   IOField "I/O field_31" at 476,376 size 58x21; FormatPattern s99999
      ProcessValue <- "AIx_DB_Flow_4_SP_SC"
   IOField "I/O field_32" at 250,358 size 58x21; FormatPattern 99999
      ProcessValue <- "AIx_DB_Flow_4_SP_HH"
   IOField "I/O field_33" at 250,378 size 58x21; FormatPattern 99999
      ProcessValue <- "AIx_DB_Flow_4_SP_H"
   IOField "I/O field_34" at 250,398 size 58x21; FormatPattern s99999
      ProcessValue <- "AIx_DB_Flow_4_SP_L"
   IOField "I/O field_35" at 250,418 size 58x21; FormatPattern s99999
      ProcessValue <- "AIx_DB_Flow_4_SP_LL"
   IOField "I/O field_36" at 550,356 size 58x21; FormatPattern 999
      ProcessValue <- "AIx_DB_Flow_4_Timers_NC_SP"
   IOField "I/O field_37" at 550,376 size 58x21; FormatPattern 999
      ProcessValue <- "AIx_DB_Flow_4_Timers_SC_SP"
   IOField "I/O field_38" at 324,358 size 58x21; FormatPattern 999
      ProcessValue <- "AIx_DB_Flow_4_Timers_HH_SP"
   IOField "I/O field_39" at 324,378 size 58x21; FormatPattern 999
      ProcessValue <- "AIx_DB_Flow_4_Timers_H_SP"
   IOField "I/O field_40" at 324,398 size 58x21; FormatPattern 999
      ProcessValue <- "AIx_DB_Flow_4_Timers_L_SP"
   IOField "I/O field_41" at 324,418 size 58x21; FormatPattern 999
      ProcessValue <- "AIx_DB_Flow_4_Timers_LL_SP"
   IOField "I/O field_42" at 586,326 size 65x25; FormatPattern s99999
      ProcessValue <- "AIx_DB_Flow_4_Signal"
   TextField "Text field_29" at 214,330 size 68x22; Text 'Уставка'
   TextField "Text field_30" at 303,330 size 79x22; Text 'Время (с)'
   Button "Button_1" at 7,5 size 96x32; TextOff 'Насосы'; Authorization "Admin"
      on Release: ActivateScreen("Dos", 0); SetTag("settings", 1)
      Appearance <- "settings"
   Button "Button_2" at 7,51 size 96x32; TextOff 'Расход-1'; Authorization "Admin"
      on Release: ActivateScreen("Flow", 0); SetTag("settings", 2)
      Appearance <- "settings"
   Button "Button_3" at 7,140 size 96x32; TextOff 'Мутность'; Authorization "Admin"
      on Release: ActivateScreen("Trans", 0); SetTag("settings", 4)
      Appearance <- "settings"
   Button "Button_5" at 7,184 size 96x32; TextOff 'DI'; Authorization "Admin"
      on Release: ActivateScreen("DI", 0); SetTag("settings", 5)
      Appearance <- "settings"
   Button "Button_6" at 7,229 size 96x32; TextOff 'DO'; Authorization "Admin"
      on Release: ActivateScreen("DO", 0); SetTag("settings", 6)
      Appearance <- "settings"
   Button "Button_4" at 7,274 size 96x32; TextOff 'PID'; Authorization "Admin"
      on Release: ActivateScreen("PID_settings", 0); SetTag("settings", 7)
      Appearance <- "settings"
   Button "Button_15" at 7,95 size 96x32; TextOff 'Расход-2'; Authorization "Admin"
      on Release: ActivateScreen("Flow_1", 0); SetTag("settings", 3)
      Appearance <- "settings"
*)

(* ===== HMI "HMI_RT_4" =====
system functions are stored by id; their names below are inferred from use
connection "HMI_Connection_2": ETHERNET, SMART_S7_1200_OMS

HMI tags "Default tag table"
   "Comm_1_DB_Mix_3_Status" : Int = PLC Comm_1_DB.Mix_3_Status AT %DB11.DBW24, 1 s
   "Comm_1_DB_Mix_2_Status" : Int = PLC Comm_1_DB.Mix_2_Status AT %DB11.DBW18, 1 s
   "Comm_1_DB_Mix_1_Status" : Int = PLC Comm_1_DB.Mix_1_Status AT %DB11.DBW12, 1 s
   "Comm_1_DB_Level" : Real = PLC Comm_1_DB.Level AT %DB11.DBD38, 1 s
   "Comm_2_DB_Level" : Real = PLC Comm_2_DB.Level AT %DB12.DBD38, 1 s
   "Comm_2_DB_Mix_1_Status" : Int = PLC Comm_2_DB.Mix_1_Status AT %DB12.DBW12, 1 s
   "Comm_2_DB_Mix_2_Status" : Int = PLC Comm_2_DB.Mix_2_Status AT %DB12.DBW18, 1 s
   "Comm_2_DB_Mix_3_Status" : Int = PLC Comm_2_DB.Mix_3_Status AT %DB12.DBW24, 1 s
   "Any_Hand" : Bool = PLC Any_Hand AT %M5.0, 1 s
   "Logick_DB_Start" : Bool = PLC Logick_DB.Start AT %DB1.DBX0.0, 1 s
   "Logick_DB_Hand" : Bool = PLC Logick_DB.Hand AT %DB1.DBX0.1, 1 s
   "Logick_DB_Use_M1" : Bool = PLC Logick_DB.Use_M1 AT %DB1.DBX0.6, 1 s
   "Logick_DB_Use_M3" : Bool = PLC Logick_DB.Use_M3 AT %DB1.DBX1.0, 1 s
   "Logick_DB_REQ_M2_1" : Bool = PLC Logick_DB.REQ_M2_1 AT %DB1.DBX1.3, 1 s
   "Logick_DB_Res_M1" : Bool = PLC Logick_DB.Res_M1 AT %DB1.DBX1.1, 1 s
   "Logick_DB_Res_M3" : Bool = PLC Logick_DB.Res_M3 AT %DB1.DBX1.2, 1 s
   "RS232_DB_Mass_1" : Real = PLC RS232_DB.Mass_1 AT %DB2.DBD0, 1 s
   "Statistics_DB_Today_1" : Real = PLC Statistics_DB.Today_1 AT %DB4.DBD40, 1 s
   "Statistics_DB_Mass_2" : Real = PLC Statistics_DB.Mass_2 AT %DB4.DBD4, 1 s
   "Statistics_DB_Mass_1" : Real = PLC Statistics_DB.Mass_1 AT %DB4.DBD0, 1 s
   "Statistics_DB_Today_2" : Real = PLC Statistics_DB.Today_2 AT %DB4.DBD44, 1 s
   "Logick_DB_Fix_1" : Bool = PLC Logick_DB.Fix_1 AT %DB1.DBX0.2, 1 s
   "Logick_DB_Fix_D_1" : Real = PLC Logick_DB.Fix_D_1 AT %DB1.DBD48, 1 s
   "Logick_DB_D_1" : Real = PLC Logick_DB.D_1 AT %DB1.DBD56, 1 s
   "Logick_DB_Fix_2" : Bool = PLC Logick_DB.Fix_2 AT %DB1.DBX0.3, 1 s
   "Logick_DB_Fix_D_2" : Real = PLC Logick_DB.Fix_D_2 AT %DB1.DBD52, 1 s
   "Logick_DB_D_2" : Real = PLC Logick_DB.D_2 AT %DB1.DBD60, 1 s
   "Comm_1_DB_Warning" : Bool = PLC Comm_1_DB.Warning AT %DB11.DBX48.2, 1 s
   "Comm_2_DB_Warning" : Bool = PLC Comm_2_DB.Warning AT %DB12.DBX48.2, 1 s
   "Logick_DB_C_1" : Real = PLC Logick_DB.C_1 AT %DB1.DBD64, 1 s
   "Logick_DB_C_2" : Real = PLC Logick_DB.C_2 AT %DB1.DBD68, 1 s
   "Statistics_DB_Zero_1" : Real = PLC Statistics_DB.Zero_1 AT %DB4.DBD64, 1 s
   "RS232_DB_Mass_2" : Real = PLC RS232_DB.Mass_2 AT %DB2.DBD4, 1 s
   "Statistics_DB_Zero_2" : Real = PLC Statistics_DB.Zero_2 AT %DB4.DBD68, 1 s
   "Statistics_DB_Last_1" : Real = PLC Statistics_DB.Last_1 AT %DB4.DBD24, 1 s
   "Statistics_DB_Delta_1" : Real = PLC Statistics_DB.Delta_1 AT %DB4.DBD32, 1 s
   "Statistics_DB_Max_D_1" : Real = PLC Statistics_DB.Max_D_1 AT %DB4.DBD16, 1 s
   "Statistics_DB_Min_D_1" : Real = PLC Statistics_DB.Min_D_1 AT %DB4.DBD8, 1 s
   "Statistics_DB_T_SP_M" : Int = PLC Statistics_DB.T.SP_M AT %DB4.DBW580, 1 s
   "Statistics_DB_T_SP_S" : Int = PLC Statistics_DB.T.SP_S AT %DB4.DBW582, 1 s
   "Sync" : Bool = PLC Sync_1 AT %M10.0, 1 s
   "Sync_2" : Bool = PLC Sync_2 AT %M10.1, 1 s
   "Statistics_DB_Delta_2" : Real = PLC Statistics_DB.Delta_2 AT %DB4.DBD36, 1 s
   "Statistics_DB_Last_2" : Real = PLC Statistics_DB.Last_2 AT %DB4.DBD28, 1 s
   "Statistics_DB_Max_D_2" : Real = PLC Statistics_DB.Max_D_2 AT %DB4.DBD20, 1 s
   "Statistics_DB_Min_D_2" : Real = PLC Statistics_DB.Min_D_2 AT %DB4.DBD12, 1 s
   "DIx_DB_Heat_4_Signal" : Bool = PLC DIx_DB.Heat_4.Signal AT %DB200.DBX122.0, 1 s
   "DIx_DB_Heat_4_Input" : Bool = PLC DIx_DB.Heat_4.Input AT %DB200.DBX120.0, 1 s
   "DIx_DB_Heat_1_Inverse" : Bool = PLC DIx_DB.Heat_1.Inverse AT %DB200.DBX64.3, 1 s
   "Any_Alm" : Bool = PLC Any_Alm AT %M6.0, 1 s
   "Statistics_DB_Today_Int" : Int = PLC Statistics_DB.Today_Int AT %DB4.DBW74, 1 s
   "Time_Save" : Bool = PLC "Time".Save AT %DB13.DBX38.0, 1 s
   "Time_Year" : UInt = PLC "Time".Year AT %DB13.DBW28, 1 s
   "Time_Month" : UInt = PLC "Time".Month AT %DB13.DBW30, 1 s
   "Time_Day" : UInt = PLC "Time".Day AT %DB13.DBW32, 1 s
   "Time_Hour" : UInt = PLC "Time".Hour AT %DB13.DBW34, 1 s
   "Time_Minutes" : UInt = PLC "Time".Minutes AT %DB13.DBW36, 1 s
   "Time_Today_YEAR" : UInt = PLC "Time".Today.YEAR AT %DB13.DBW0, 1 s
   "Time_Today_MONTH" : USInt = PLC "Time".Today.MONTH AT %DB13.DBB2, 1 s
   "Time_Today_DAY" : USInt = PLC "Time".Today.DAY AT %DB13.DBB3, 1 s
   "Time_Today_WEEKDAY" : USInt = PLC "Time".Today.WEEKDAY AT %DB13.DBB4, 1 s
   "Time_Today_HOUR" : USInt = PLC "Time".Today.HOUR AT %DB13.DBB5, 1 s
   "Time_Today_MINUTE" : USInt = PLC "Time".Today.MINUTE AT %DB13.DBB6, 1 s
   "Reset_All" : Bool = PLC Reset_All AT %M3.1, 1 s
   "Logick_DB_Low_REQ" : Bool = PLC Logick_DB.Low_REQ AT %DB1.DBX2.0, 1 s
   "Logick_DB_Low_view" : Bool = PLC Logick_DB.Low_view AT %DB1.DBX2.2, 1 s
   "Logick_DB_Low_SP_M" : Int = PLC Logick_DB.Low.SP_M AT %DB1.DBW72, 1 s
   "Logick_DB_Low_CMD" : Bool = PLC Logick_DB.Low_CMD AT %DB1.DBX2.1, 1 s
   "Logick_DB_Max_SP" : Real = PLC Logick_DB.Max_SP AT %DB1.DBD36, 1 s
   "Logick_DB_Min_SP" : Real = PLC Logick_DB.Min_SP AT %DB1.DBD32, 1 s
   "Logick_DB_Low_use" : Bool = PLC Logick_DB.Low_use AT %DB1.DBX1.7, 1 s

HMI tags "HMI"
   "settings" : Int, internal

HMI tags "xDI"
   "DIx_DB_M1_QF_Input" : Bool = PLC DIx_DB.M1_QF.Input AT %DB200.DBX0.0, 1 s
   "DIx_DB_M1_QF_Signal" : Bool = PLC DIx_DB.M1_QF.Signal AT %DB200.DBX2.0, 1 s
   "DIx_DB_M1_QF_Hand" : Bool = PLC DIx_DB.M1_QF.Hand AT %DB200.DBX4.0, 1 s
   "DIx_DB_M1_QF_Start_M" : Bool = PLC DIx_DB.M1_QF.Start_M AT %DB200.DBX4.1, 1 s
   "DIx_DB_M1_QF_Inverse" : Bool = PLC DIx_DB.M1_QF.Inverse AT %DB200.DBX4.3, 1 s
   "DIx_DB_M1_QF_Filter_On_SP" : Int = PLC DIx_DB.M1_QF.Filter_On.SP AT %DB200.DBW6, 1 s
   "DIx_DB_M1_QF_Filter_Off_SP" : Int = PLC DIx_DB.M1_QF.Filter_Off.SP AT %DB200.DBW12, 1 s
   "DIx_DB_M2_QF_Input" : Bool = PLC DIx_DB.M2_QF.Input AT %DB200.DBX20.0, 1 s
   "DIx_DB_M2_QF_Signal" : Bool = PLC DIx_DB.M2_QF.Signal AT %DB200.DBX22.0, 1 s
   "DIx_DB_M2_QF_Hand" : Bool = PLC DIx_DB.M2_QF.Hand AT %DB200.DBX24.0, 1 s
   "DIx_DB_M2_QF_Start_M" : Bool = PLC DIx_DB.M2_QF.Start_M AT %DB200.DBX24.1, 1 s
   "DIx_DB_M2_QF_Inverse" : Bool = PLC DIx_DB.M2_QF.Inverse AT %DB200.DBX24.3, 1 s
   "DIx_DB_M2_QF_Filter_On_SP" : Int = PLC DIx_DB.M2_QF.Filter_On.SP AT %DB200.DBW26, 1 s
   "DIx_DB_M2_QF_Filter_Off_SP" : Int = PLC DIx_DB.M2_QF.Filter_Off.SP AT %DB200.DBW32, 1 s
   "DIx_DB_M3_QF_Input" : Bool = PLC DIx_DB.M3_QF.Input AT %DB200.DBX40.0, 1 s
   "DIx_DB_M3_QF_Signal" : Bool = PLC DIx_DB.M3_QF.Signal AT %DB200.DBX42.0, 1 s
   "DIx_DB_M3_QF_Hand" : Bool = PLC DIx_DB.M3_QF.Hand AT %DB200.DBX44.0, 1 s
   "DIx_DB_M3_QF_Start_M" : Bool = PLC DIx_DB.M3_QF.Start_M AT %DB200.DBX44.1, 1 s
   "DIx_DB_M3_QF_Inverse" : Bool = PLC DIx_DB.M3_QF.Inverse AT %DB200.DBX44.3, 1 s
   "DIx_DB_M3_QF_Filter_On_SP" : Int = PLC DIx_DB.M3_QF.Filter_On.SP AT %DB200.DBW46, 1 s
   "DIx_DB_M3_QF_Filter_Off_SP" : Int = PLC DIx_DB.M3_QF.Filter_Off.SP AT %DB200.DBW52, 1 s
   "DIx_DB_Heat_1_Input" : Bool = PLC DIx_DB.Heat_1.Input AT %DB200.DBX60.0, 1 s
   "DIx_DB_Heat_1_Signal" : Bool = PLC DIx_DB.Heat_1.Signal AT %DB200.DBX62.0, 1 s
   "DIx_DB_Heat_1_Hand" : Bool = PLC DIx_DB.Heat_1.Hand AT %DB200.DBX64.0, 1 s
   "DIx_DB_Heat_1_Start_M" : Bool = PLC DIx_DB.Heat_1.Start_M AT %DB200.DBX64.1, 1 s
   "DIx_DB_Heat_1_Filter_On_SP" : Int = PLC DIx_DB.Heat_1.Filter_On.SP AT %DB200.DBW66, 1 s
   "DIx_DB_Heat_1_Filter_Off_SP" : Int = PLC DIx_DB.Heat_1.Filter_Off.SP AT %DB200.DBW72, 1 s
   "DIx_DB_Heat_2_Filter_Off_SP" : Int = PLC DIx_DB.Heat_2.Filter_Off.SP AT %DB200.DBW92, 1 s
   "DIx_DB_Heat_2_Filter_On_SP" : Int = PLC DIx_DB.Heat_2.Filter_On.SP AT %DB200.DBW86, 1 s
   "DIx_DB_Heat_2_Inverse" : Bool = PLC DIx_DB.Heat_2.Inverse AT %DB200.DBX84.3, 1 s
   "DIx_DB_Heat_2_Start_M" : Bool = PLC DIx_DB.Heat_2.Start_M AT %DB200.DBX84.1, 1 s
   "DIx_DB_Heat_2_Hand" : Bool = PLC DIx_DB.Heat_2.Hand AT %DB200.DBX84.0, 1 s
   "DIx_DB_Heat_2_Signal" : Bool = PLC DIx_DB.Heat_2.Signal AT %DB200.DBX82.0, 1 s
   "DIx_DB_Heat_2_Input" : Bool = PLC DIx_DB.Heat_2.Input AT %DB200.DBX80.0, 1 s
   "DIx_DB_Heat_3_Input" : Bool = PLC DIx_DB.Heat_3.Input AT %DB200.DBX100.0, 1 s
   "DIx_DB_Heat_3_Signal" : Bool = PLC DIx_DB.Heat_3.Signal AT %DB200.DBX102.0, 1 s
   "DIx_DB_Heat_3_Hand" : Bool = PLC DIx_DB.Heat_3.Hand AT %DB200.DBX104.0, 1 s
   "DIx_DB_Heat_3_Start_M" : Bool = PLC DIx_DB.Heat_3.Start_M AT %DB200.DBX104.1, 1 s
   "DIx_DB_Heat_3_Inverse" : Bool = PLC DIx_DB.Heat_3.Inverse AT %DB200.DBX104.3, 1 s
   "DIx_DB_Heat_3_Filter_Off_SP" : Int = PLC DIx_DB.Heat_3.Filter_Off.SP AT %DB200.DBW112, 1 s
   "DIx_DB_Heat_3_Filter_On_SP" : Int = PLC DIx_DB.Heat_3.Filter_On.SP AT %DB200.DBW106, 1 s
   "DIx_DB_AllBlock_Input" : Bool = PLC DIx_DB.AllBlock.Input AT %DB200.DBX140.0, 1 s
   "DIx_DB_AllBlock_Signal" : Bool = PLC DIx_DB.AllBlock.Signal AT %DB200.DBX142.0, 1 s
   "DIx_DB_AllBlock_Hand" : Bool = PLC DIx_DB.AllBlock.Hand AT %DB200.DBX144.0, 1 s
   "DIx_DB_AllBlock_Start_M" : Bool = PLC DIx_DB.AllBlock.Start_M AT %DB200.DBX144.1, 1 s
   "DIx_DB_AllBlock_Inverse" : Bool = PLC DIx_DB.AllBlock.Inverse AT %DB200.DBX144.3, 1 s
   "DIx_DB_AllBlock_Filter_On_SP" : Int = PLC DIx_DB.AllBlock.Filter_On.SP AT %DB200.DBW146, 1 s
   "DIx_DB_AllBlock_Filter_Off_SP" : Int = PLC DIx_DB.AllBlock.Filter_Off.SP AT %DB200.DBW152, 1 s
   "DIx_DB_Mass_1_Input" : Bool = PLC DIx_DB.Mass_1.Input AT %DB200.DBX160.0, 1 s
   "DIx_DB_Mass_1_Signal" : Bool = PLC DIx_DB.Mass_1.Signal AT %DB200.DBX162.0, 1 s
   "DIx_DB_Mass_1_Hand" : Bool = PLC DIx_DB.Mass_1.Hand AT %DB200.DBX164.0, 1 s
   "DIx_DB_Mass_1_Start_M" : Bool = PLC DIx_DB.Mass_1.Start_M AT %DB200.DBX164.1, 1 s
   "DIx_DB_Mass_1_Inverse" : Bool = PLC DIx_DB.Mass_1.Inverse AT %DB200.DBX164.3, 1 s
   "DIx_DB_Mass_1_Filter_On_SP" : Int = PLC DIx_DB.Mass_1.Filter_On.SP AT %DB200.DBW166, 1 s
   "DIx_DB_Mass_1_Filter_Off_SP" : Int = PLC DIx_DB.Mass_1.Filter_Off.SP AT %DB200.DBW172, 1 s
   "DIx_DB_Mass_2_Input" : Bool = PLC DIx_DB.Mass_2.Input AT %DB200.DBX180.0, 1 s
   "DIx_DB_Mass_2_Signal" : Bool = PLC DIx_DB.Mass_2.Signal AT %DB200.DBX182.0, 1 s
   "DIx_DB_Mass_2_Hand" : Bool = PLC DIx_DB.Mass_2.Hand AT %DB200.DBX184.0, 1 s
   "DIx_DB_Mass_2_Start_M" : Bool = PLC DIx_DB.Mass_2.Start_M AT %DB200.DBX184.1, 1 s
   "DIx_DB_Mass_2_Inverse" : Bool = PLC DIx_DB.Mass_2.Inverse AT %DB200.DBX184.3, 1 s
   "DIx_DB_Mass_2_Filter_On_SP" : Int = PLC DIx_DB.Mass_2.Filter_On.SP AT %DB200.DBW186, 1 s
   "DIx_DB_Mass_2_Filter_Off_SP" : Int = PLC DIx_DB.Mass_2.Filter_Off.SP AT %DB200.DBW192, 1 s
   "DIx_DB_Heat_4_Hand" : Bool = PLC DIx_DB.Heat_4.Hand AT %DB200.DBX124.0, 1 s
   "DIx_DB_Heat_4_Start_M" : Bool = PLC DIx_DB.Heat_4.Start_M AT %DB200.DBX124.1, 1 s
   "DIx_DB_Heat_4_Inverse" : Bool = PLC DIx_DB.Heat_4.Inverse AT %DB200.DBX124.3, 1 s
   "DIx_DB_Heat_4_Filter_On_SP" : Int = PLC DIx_DB.Heat_4.Filter_On.SP AT %DB200.DBW126, 1 s
   "DIx_DB_Heat_4_Filter_Off_SP" : Int = PLC DIx_DB.Heat_4.Filter_Off.SP AT %DB200.DBW132, 1 s

HMI tags "xDO"
   "DOx_DB_M1_CMD_Start_A" : Bool = PLC DOx_DB.M1_CMD.Start_A AT %DB201.DBX0.0, 1 s
   "DOx_DB_M1_CMD_Q" : Bool = PLC DOx_DB.M1_CMD.Q AT %DB201.DBX0.2, 1 s
   "DOx_DB_M1_CMD_Hand" : Bool = PLC DOx_DB.M1_CMD.Hand AT %DB201.DBX2.0, 1 s
   "DOx_DB_M1_CMD_Start_M" : Bool = PLC DOx_DB.M1_CMD.Start_M AT %DB201.DBX2.1, 1 s
   "DOx_DB_M1_CMD_Simulation" : Bool = PLC DOx_DB.M1_CMD.Simulation AT %DB201.DBX2.2, 1 s
   "DOx_DB_M1_CMD_Inverse" : Bool = PLC DOx_DB.M1_CMD.Inverse AT %DB201.DBX2.3, 1 s
   "DOx_DB_M2_CMD_Start_A" : Bool = PLC DOx_DB.M2_CMD.Start_A AT %DB201.DBX10.0, 1 s
   "DOx_DB_M2_CMD_Q" : Bool = PLC DOx_DB.M2_CMD.Q AT %DB201.DBX10.2, 1 s
   "DOx_DB_M2_CMD_Hand" : Bool = PLC DOx_DB.M2_CMD.Hand AT %DB201.DBX12.0, 1 s
   "DOx_DB_M2_CMD_Start_M" : Bool = PLC DOx_DB.M2_CMD.Start_M AT %DB201.DBX12.1, 1 s
   "DOx_DB_M2_CMD_Simulation" : Bool = PLC DOx_DB.M2_CMD.Simulation AT %DB201.DBX12.2, 1 s
   "DOx_DB_M2_CMD_Inverse" : Bool = PLC DOx_DB.M2_CMD.Inverse AT %DB201.DBX12.3, 1 s
   "DOx_DB_M3_CMD_Start_A" : Bool = PLC DOx_DB.M3_CMD.Start_A AT %DB201.DBX20.0, 1 s
   "DOx_DB_M3_CMD_Q" : Bool = PLC DOx_DB.M3_CMD.Q AT %DB201.DBX20.2, 1 s
   "DOx_DB_M3_CMD_Hand" : Bool = PLC DOx_DB.M3_CMD.Hand AT %DB201.DBX22.0, 1 s
   "DOx_DB_M3_CMD_Start_M" : Bool = PLC DOx_DB.M3_CMD.Start_M AT %DB201.DBX22.1, 1 s
   "DOx_DB_M3_CMD_Simulation" : Bool = PLC DOx_DB.M3_CMD.Simulation AT %DB201.DBX22.2, 1 s
   "DOx_DB_M3_CMD_Inverse" : Bool = PLC DOx_DB.M3_CMD.Inverse AT %DB201.DBX22.3, 1 s
   "DOx_DB_LED_Error_1_Start_A" : Bool = PLC DOx_DB.LED_Error_1.Start_A AT %DB201.DBX30.0, 1 s
   "DOx_DB_LED_Error_1_Q" : Bool = PLC DOx_DB.LED_Error_1.Q AT %DB201.DBX30.2, 1 s
   "DOx_DB_LED_Error_1_Hand" : Bool = PLC DOx_DB.LED_Error_1.Hand AT %DB201.DBX32.0, 1 s
   "DOx_DB_LED_Error_1_Simulation" : Bool = PLC DOx_DB.LED_Error_1.Simulation AT %DB201.DBX32.2, 1 s
   "DOx_DB_LED_Error_1_Start_M" : Bool = PLC DOx_DB.LED_Error_1.Start_M AT %DB201.DBX32.1, 1 s
   "DOx_DB_LED_Error_1_Inverse" : Bool = PLC DOx_DB.LED_Error_1.Inverse AT %DB201.DBX32.3, 1 s
   "DOx_DB_LED_Error_2_Start_A" : Bool = PLC DOx_DB.LED_Error_2.Start_A AT %DB201.DBX40.0, 1 s
   "DOx_DB_LED_Error_2_Q" : Bool = PLC DOx_DB.LED_Error_2.Q AT %DB201.DBX40.2, 1 s
   "DOx_DB_LED_Error_2_Hand" : Bool = PLC DOx_DB.LED_Error_2.Hand AT %DB201.DBX42.0, 1 s
   "DOx_DB_LED_Error_2_Start_M" : Bool = PLC DOx_DB.LED_Error_2.Start_M AT %DB201.DBX42.1, 1 s
   "DOx_DB_LED_Error_2_Simulation" : Bool = PLC DOx_DB.LED_Error_2.Simulation AT %DB201.DBX42.2, 1 s
   "DOx_DB_LED_Error_2_Inverse" : Bool = PLC DOx_DB.LED_Error_2.Inverse AT %DB201.DBX42.3, 1 s
   "DOx_DB_LED_Alarm_Start_A" : Bool = PLC DOx_DB.LED_Alarm.Start_A AT %DB201.DBX50.0, 1 s
   "DOx_DB_LED_Alarm_Q" : Bool = PLC DOx_DB.LED_Alarm.Q AT %DB201.DBX50.2, 1 s
   "DOx_DB_LED_Alarm_Hand" : Bool = PLC DOx_DB.LED_Alarm.Hand AT %DB201.DBX52.0, 1 s
   "DOx_DB_LED_Alarm_Start_M" : Bool = PLC DOx_DB.LED_Alarm.Start_M AT %DB201.DBX52.1, 1 s
   "DOx_DB_LED_Alarm_Simulation" : Bool = PLC DOx_DB.LED_Alarm.Simulation AT %DB201.DBX52.2, 1 s
   "DOx_DB_LED_Alarm_Inverse" : Bool = PLC DOx_DB.LED_Alarm.Inverse AT %DB201.DBX52.3, 1 s
   "DOx_DB_LED_M1_Alarm_Start_A" : Bool = PLC DOx_DB.LED_M1_Alarm.Start_A AT %DB201.DBX60.0, 1 s
   "DOx_DB_LED_M1_Alarm_Q" : Bool = PLC DOx_DB.LED_M1_Alarm.Q AT %DB201.DBX60.2, 1 s
   "DOx_DB_LED_M1_Alarm_Hand" : Bool = PLC DOx_DB.LED_M1_Alarm.Hand AT %DB201.DBX62.0, 1 s
   "DOx_DB_LED_M1_Alarm_Start_M" : Bool = PLC DOx_DB.LED_M1_Alarm.Start_M AT %DB201.DBX62.1, 1 s
   "DOx_DB_LED_M1_Alarm_Simulation" : Bool = PLC DOx_DB.LED_M1_Alarm.Simulation AT %DB201.DBX62.2, 1 s
   "DOx_DB_LED_M1_Alarm_Inverse" : Bool = PLC DOx_DB.LED_M1_Alarm.Inverse AT %DB201.DBX62.3, 1 s
   "DOx_DB_LED_M2_Alarm_Start_A" : Bool = PLC DOx_DB.LED_M2_Alarm.Start_A AT %DB201.DBX70.0, 1 s
   "DOx_DB_LED_M2_Alarm_Q" : Bool = PLC DOx_DB.LED_M2_Alarm.Q AT %DB201.DBX70.2, 1 s
   "DOx_DB_LED_M2_Alarm_Hand" : Bool = PLC DOx_DB.LED_M2_Alarm.Hand AT %DB201.DBX72.0, 1 s
   "DOx_DB_LED_M2_Alarm_Start_M" : Bool = PLC DOx_DB.LED_M2_Alarm.Start_M AT %DB201.DBX72.1, 1 s
   "DOx_DB_LED_M2_Alarm_Simulation" : Bool = PLC DOx_DB.LED_M2_Alarm.Simulation AT %DB201.DBX72.2, 1 s
   "DOx_DB_LED_M2_Alarm_Inverse" : Bool = PLC DOx_DB.LED_M2_Alarm.Inverse AT %DB201.DBX72.3, 1 s
   "DOx_DB_LED_M3_Alarm_Start_A" : Bool = PLC DOx_DB.LED_M3_Alarm.Start_A AT %DB201.DBX80.0, 1 s
   "DOx_DB_LED_M3_Alarm_Q" : Bool = PLC DOx_DB.LED_M3_Alarm.Q AT %DB201.DBX80.2, 1 s
   "DOx_DB_LED_M3_Alarm_Hand" : Bool = PLC DOx_DB.LED_M3_Alarm.Hand AT %DB201.DBX82.0, 1 s
   "DOx_DB_LED_M3_Alarm_Start_M" : Bool = PLC DOx_DB.LED_M3_Alarm.Start_M AT %DB201.DBX82.1, 1 s
   "DOx_DB_LED_M3_Alarm_Simulation" : Bool = PLC DOx_DB.LED_M3_Alarm.Simulation AT %DB201.DBX82.2, 1 s
   "DOx_DB_LED_M3_Alarm_Inverse" : Bool = PLC DOx_DB.LED_M3_Alarm.Inverse AT %DB201.DBX82.3, 1 s

HMI tags "xAI"
   "AIx_DB_Flow_1_Signal" : Int = PLC AIx_DB.Flow_1.Signal AT %DB202.DBW0, 1 s
   "AIx_DB_Flow_1_Result" : Real = PLC AIx_DB.Flow_1.Result AT %DB202.DBD6, 1 s
   "AIx_DB_Flow_1_CMD_Start_A" : Bool = PLC AIx_DB.Flow_1.CMD.Start_A AT %DB202.DBX10.1, 1 s
   "AIx_DB_Flow_1_CMD_Hand" : Bool = PLC AIx_DB.Flow_1.CMD.Hand AT %DB202.DBX10.0, 1 s
   "AIx_DB_Flow_1_Use_RTD" : Bool = PLC AIx_DB.Flow_1.Use.RTD AT %DB202.DBX16.0, 1 s
   "AIx_DB_Flow_1_Use_Filter" : Bool = PLC AIx_DB.Flow_1.Use.Filter AT %DB202.DBX16.1, 1 s
   "AIx_DB_Flow_1_RTD_c" : Real = PLC AIx_DB.Flow_1.RTD_c AT %DB202.DBD30, 1 s
   "AIx_DB_Flow_1_Calibration" : Real = PLC AIx_DB.Flow_1.Calibration AT %DB202.DBD34, 1 s
   "AIx_DB_Flow_1_Converter_Min_In" : Real = PLC AIx_DB.Flow_1.Converter.Min_In AT %DB202.DBD60, 1 s
   "AIx_DB_Flow_1_Converter_Max_In" : Real = PLC AIx_DB.Flow_1.Converter.Max_In AT %DB202.DBD64, 1 s
   "AIx_DB_Flow_1_Converter_Min_Out" : Real = PLC AIx_DB.Flow_1.Converter.Min_Out AT %DB202.DBD68, 1 s
   "AIx_DB_Flow_1_Converter_Max_Out" : Real = PLC AIx_DB.Flow_1.Converter.Max_Out AT %DB202.DBD72, 1 s
   "AIx_DB_Flow_1_Filter_SP" : Real = PLC AIx_DB.Flow_1.Filter.SP AT %DB202.DBD38, 1 s
   "AIx_DB_Flow_1_SP_NC" : Real = PLC AIx_DB.Flow_1.SP.NC AT %DB202.DBD76, 1 s
   "AIx_DB_Flow_1_SP_SC" : Real = PLC AIx_DB.Flow_1.SP.SC AT %DB202.DBD80, 1 s
   "AIx_DB_Flow_1_SP_HH" : Real = PLC AIx_DB.Flow_1.SP.HH AT %DB202.DBD84, 1 s
   "AIx_DB_Flow_1_SP_H" : Real = PLC AIx_DB.Flow_1.SP.H AT %DB202.DBD88, 1 s
   "AIx_DB_Flow_1_SP_L" : Real = PLC AIx_DB.Flow_1.SP.L AT %DB202.DBD92, 1 s
   "AIx_DB_Flow_1_SP_LL" : Real = PLC AIx_DB.Flow_1.SP.LL AT %DB202.DBD96, 1 s
   "AIx_DB_Flow_1_Alarm" : Word = PLC AIx_DB.Flow_1.Alarm AT %DB202.DBW138, 1 s
   "AIx_DB_Flow_1_Timers_NC_SP" : Int = PLC AIx_DB.Flow_1.Timers.NC.SP AT %DB202.DBW100, 1 s
   "AIx_DB_Flow_1_Timers_SC_SP" : Int = PLC AIx_DB.Flow_1.Timers.SC.SP AT %DB202.DBW106, 1 s
   "AIx_DB_Flow_1_Timers_HH_SP" : Int = PLC AIx_DB.Flow_1.Timers.HH.SP AT %DB202.DBW112, 1 s
   "AIx_DB_Flow_1_Timers_H_SP" : Int = PLC AIx_DB.Flow_1.Timers.H.SP AT %DB202.DBW118, 1 s
   "AIx_DB_Flow_1_Timers_L_SP" : Int = PLC AIx_DB.Flow_1.Timers.L.SP AT %DB202.DBW124, 1 s
   "AIx_DB_Flow_1_Timers_LL_SP" : Int = PLC AIx_DB.Flow_1.Timers.LL.SP AT %DB202.DBW130, 1 s
   "AIx_DB_Flow_2_Signal" : Int = PLC AIx_DB.Flow_2.Signal AT %DB202.DBW140, 1 s
   "AIx_DB_Flow_2_Result" : Real = PLC AIx_DB.Flow_2.Result AT %DB202.DBD146, 1 s
   "AIx_DB_Flow_2_CMD_Start_A" : Bool = PLC AIx_DB.Flow_2.CMD.Start_A AT %DB202.DBX150.1, 1 s
   "AIx_DB_Flow_2_CMD_Hand" : Bool = PLC AIx_DB.Flow_2.CMD.Hand AT %DB202.DBX150.0, 1 s
   "AIx_DB_Flow_2_Use_RTD" : Bool = PLC AIx_DB.Flow_2.Use.RTD AT %DB202.DBX156.0, 1 s
   "AIx_DB_Flow_2_Use_Filter" : Bool = PLC AIx_DB.Flow_2.Use.Filter AT %DB202.DBX156.1, 1 s
   "AIx_DB_Flow_2_RTD_c" : Real = PLC AIx_DB.Flow_2.RTD_c AT %DB202.DBD170, 1 s
   "AIx_DB_Flow_2_Calibration" : Real = PLC AIx_DB.Flow_2.Calibration AT %DB202.DBD174, 1 s
   "AIx_DB_Flow_2_Converter_Min_In" : Real = PLC AIx_DB.Flow_2.Converter.Min_In AT %DB202.DBD200, 1 s
   "AIx_DB_Flow_2_Converter_Max_In" : Real = PLC AIx_DB.Flow_2.Converter.Max_In AT %DB202.DBD204, 1 s
   "AIx_DB_Flow_2_Converter_Min_Out" : Real = PLC AIx_DB.Flow_2.Converter.Min_Out AT %DB202.DBD208, 1 s
   "AIx_DB_Flow_2_Converter_Max_Out" : Real = PLC AIx_DB.Flow_2.Converter.Max_Out AT %DB202.DBD212, 1 s
   "AIx_DB_Flow_2_Filter_SP" : Real = PLC AIx_DB.Flow_2.Filter.SP AT %DB202.DBD178, 1 s
   "AIx_DB_Flow_2_SP_NC" : Real = PLC AIx_DB.Flow_2.SP.NC AT %DB202.DBD216, 1 s
   "AIx_DB_Flow_2_SP_SC" : Real = PLC AIx_DB.Flow_2.SP.SC AT %DB202.DBD220, 1 s
   "AIx_DB_Flow_2_SP_HH" : Real = PLC AIx_DB.Flow_2.SP.HH AT %DB202.DBD224, 1 s
   "AIx_DB_Flow_2_SP_H" : Real = PLC AIx_DB.Flow_2.SP.H AT %DB202.DBD228, 1 s
   "AIx_DB_Flow_2_SP_L" : Real = PLC AIx_DB.Flow_2.SP.L AT %DB202.DBD232, 1 s
   "AIx_DB_Flow_2_SP_LL" : Real = PLC AIx_DB.Flow_2.SP.LL AT %DB202.DBD236, 1 s
   "AIx_DB_Flow_2_Alarm" : Word = PLC AIx_DB.Flow_2.Alarm AT %DB202.DBW278, 1 s
   "AIx_DB_Flow_2_Timers_NC_SP" : Int = PLC AIx_DB.Flow_2.Timers.NC.SP AT %DB202.DBW240, 1 s
   "AIx_DB_Flow_2_Timers_SC_SP" : Int = PLC AIx_DB.Flow_2.Timers.SC.SP AT %DB202.DBW246, 1 s
   "AIx_DB_Flow_2_Timers_HH_SP" : Int = PLC AIx_DB.Flow_2.Timers.HH.SP AT %DB202.DBW252, 1 s
   "AIx_DB_Flow_2_Timers_H_SP" : Int = PLC AIx_DB.Flow_2.Timers.H.SP AT %DB202.DBW258, 1 s
   "AIx_DB_Flow_2_Timers_L_SP" : Int = PLC AIx_DB.Flow_2.Timers.L.SP AT %DB202.DBW264, 1 s
   "AIx_DB_Flow_2_Timers_LL_SP" : Int = PLC AIx_DB.Flow_2.Timers.LL.SP AT %DB202.DBW270, 1 s
   "AIx_DB_Trans_1_Signal" : Int = PLC AIx_DB.Trans_1.Signal AT %DB202.DBW280, 1 s
   "AIx_DB_Trans_1_Result" : Real = PLC AIx_DB.Trans_1.Result AT %DB202.DBD286, 1 s
   "AIx_DB_Trans_1_CMD_Start_A" : Bool = PLC AIx_DB.Trans_1.CMD.Start_A AT %DB202.DBX290.1, 1 s
   "AIx_DB_Trans_1_CMD_Hand" : Bool = PLC AIx_DB.Trans_1.CMD.Hand AT %DB202.DBX290.0, 1 s
   "AIx_DB_Trans_1_Use_RTD" : Bool = PLC AIx_DB.Trans_1.Use.RTD AT %DB202.DBX296.0, 1 s
   "AIx_DB_Trans_1_Use_Filter" : Bool = PLC AIx_DB.Trans_1.Use.Filter AT %DB202.DBX296.1, 1 s
   "AIx_DB_Trans_1_RTD_c" : Real = PLC AIx_DB.Trans_1.RTD_c AT %DB202.DBD310, 1 s
   "AIx_DB_Trans_1_Calibration" : Real = PLC AIx_DB.Trans_1.Calibration AT %DB202.DBD314, 1 s
   "AIx_DB_Trans_1_Converter_Min_In" : Real = PLC AIx_DB.Trans_1.Converter.Min_In AT %DB202.DBD340, 1 s
   "AIx_DB_Trans_1_Converter_Max_In" : Real = PLC AIx_DB.Trans_1.Converter.Max_In AT %DB202.DBD344, 1 s
   "AIx_DB_Trans_1_Converter_Min_Out" : Real = PLC AIx_DB.Trans_1.Converter.Min_Out AT %DB202.DBD348, 1 s
   "AIx_DB_Trans_1_Converter_Max_Out" : Real = PLC AIx_DB.Trans_1.Converter.Max_Out AT %DB202.DBD352, 1 s
   "AIx_DB_Trans_1_Filter_SP" : Real = PLC AIx_DB.Trans_1.Filter.SP AT %DB202.DBD318, 1 s
   "AIx_DB_Trans_1_SP_NC" : Real = PLC AIx_DB.Trans_1.SP.NC AT %DB202.DBD356, 1 s
   "AIx_DB_Trans_1_SP_SC" : Real = PLC AIx_DB.Trans_1.SP.SC AT %DB202.DBD360, 1 s
   "AIx_DB_Trans_1_SP_HH" : Real = PLC AIx_DB.Trans_1.SP.HH AT %DB202.DBD364, 1 s
   "AIx_DB_Trans_1_SP_H" : Real = PLC AIx_DB.Trans_1.SP.H AT %DB202.DBD368, 1 s
   "AIx_DB_Trans_1_SP_L" : Real = PLC AIx_DB.Trans_1.SP.L AT %DB202.DBD372, 1 s
   "AIx_DB_Trans_1_SP_LL" : Real = PLC AIx_DB.Trans_1.SP.LL AT %DB202.DBD376, 1 s
   "AIx_DB_Trans_1_Alarm" : Word = PLC AIx_DB.Trans_1.Alarm AT %DB202.DBW418, 1 s
   "AIx_DB_Trans_1_Timers_NC_SP" : Int = PLC AIx_DB.Trans_1.Timers.NC.SP AT %DB202.DBW380, 1 s
   "AIx_DB_Trans_1_Timers_SC_SP" : Int = PLC AIx_DB.Trans_1.Timers.SC.SP AT %DB202.DBW386, 1 s
   "AIx_DB_Trans_1_Timers_HH_SP" : Int = PLC AIx_DB.Trans_1.Timers.HH.SP AT %DB202.DBW392, 1 s
   "AIx_DB_Trans_1_Timers_H_SP" : Int = PLC AIx_DB.Trans_1.Timers.H.SP AT %DB202.DBW398, 1 s
   "AIx_DB_Trans_1_Timers_L_SP" : Int = PLC AIx_DB.Trans_1.Timers.L.SP AT %DB202.DBW404, 1 s
   "AIx_DB_Trans_1_Timers_LL_SP" : Int = PLC AIx_DB.Trans_1.Timers.LL.SP AT %DB202.DBW410, 1 s
   "AIx_DB_Trans_2_Signal" : Int = PLC AIx_DB.Trans_2.Signal AT %DB202.DBW420, 1 s
   "AIx_DB_Trans_2_Result" : Real = PLC AIx_DB.Trans_2.Result AT %DB202.DBD426, 1 s
   "AIx_DB_Trans_2_CMD_Start_A" : Bool = PLC AIx_DB.Trans_2.CMD.Start_A AT %DB202.DBX430.1, 1 s
   "AIx_DB_Trans_2_CMD_Hand" : Bool = PLC AIx_DB.Trans_2.CMD.Hand AT %DB202.DBX430.0, 1 s
   "AIx_DB_Trans_2_Use_RTD" : Bool = PLC AIx_DB.Trans_2.Use.RTD AT %DB202.DBX436.0, 1 s
   "AIx_DB_Trans_2_Use_Filter" : Bool = PLC AIx_DB.Trans_2.Use.Filter AT %DB202.DBX436.1, 1 s
   "AIx_DB_Trans_2_RTD_c" : Real = PLC AIx_DB.Trans_2.RTD_c AT %DB202.DBD450, 1 s
   "AIx_DB_Trans_2_Calibration" : Real = PLC AIx_DB.Trans_2.Calibration AT %DB202.DBD454, 1 s
   "AIx_DB_Trans_2_Converter_Min_In" : Real = PLC AIx_DB.Trans_2.Converter.Min_In AT %DB202.DBD480, 1 s
   "AIx_DB_Trans_2_Converter_Max_In" : Real = PLC AIx_DB.Trans_2.Converter.Max_In AT %DB202.DBD484, 1 s
   "AIx_DB_Trans_2_Converter_Min_Out" : Real = PLC AIx_DB.Trans_2.Converter.Min_Out AT %DB202.DBD488, 1 s
   "AIx_DB_Trans_2_Converter_Max_Out" : Real = PLC AIx_DB.Trans_2.Converter.Max_Out AT %DB202.DBD492, 1 s
   "AIx_DB_Trans_2_Filter_SP" : Real = PLC AIx_DB.Trans_2.Filter.SP AT %DB202.DBD458, 1 s
   "AIx_DB_Trans_2_SP_NC" : Real = PLC AIx_DB.Trans_2.SP.NC AT %DB202.DBD496, 1 s
   "AIx_DB_Trans_2_SP_SC" : Real = PLC AIx_DB.Trans_2.SP.SC AT %DB202.DBD500, 1 s
   "AIx_DB_Trans_2_SP_HH" : Real = PLC AIx_DB.Trans_2.SP.HH AT %DB202.DBD504, 1 s
   "AIx_DB_Trans_2_SP_H" : Real = PLC AIx_DB.Trans_2.SP.H AT %DB202.DBD508, 1 s
   "AIx_DB_Trans_2_SP_L" : Real = PLC AIx_DB.Trans_2.SP.L AT %DB202.DBD512, 1 s
   "AIx_DB_Trans_2_SP_LL" : Real = PLC AIx_DB.Trans_2.SP.LL AT %DB202.DBD516, 1 s
   "AIx_DB_Trans_2_Alarm" : Word = PLC AIx_DB.Trans_2.Alarm AT %DB202.DBW558, 1 s
   "AIx_DB_Trans_2_Timers_NC_SP" : Int = PLC AIx_DB.Trans_2.Timers.NC.SP AT %DB202.DBW520, 1 s
   "AIx_DB_Trans_2_Timers_SC_SP" : Int = PLC AIx_DB.Trans_2.Timers.SC.SP AT %DB202.DBW526, 1 s
   "AIx_DB_Trans_2_Timers_HH_SP" : Int = PLC AIx_DB.Trans_2.Timers.HH.SP AT %DB202.DBW532, 1 s
   "AIx_DB_Trans_2_Timers_H_SP" : Int = PLC AIx_DB.Trans_2.Timers.H.SP AT %DB202.DBW538, 1 s
   "AIx_DB_Trans_2_Timers_L_SP" : Int = PLC AIx_DB.Trans_2.Timers.L.SP AT %DB202.DBW544, 1 s
   "AIx_DB_Trans_2_Timers_LL_SP" : Int = PLC AIx_DB.Trans_2.Timers.LL.SP AT %DB202.DBW550, 1 s
